
         A     "T_Highpressure_MH02";
         =     "DB123_MH_IO_Signals".MH[2].IN.MH_HP_Circ_MH;
         A     "T_Start_MH02";
         =     "DB123_MH_IO_Signals".MH[2].IN.MH_Start;
         A     "T_Stop_MH02";
         =     "DB123_MH_IO_Signals".MH[2].IN.MH_Stop;
         A     "T_CP_forward_MH02";
         =     "DB123_MH_IO_Signals".MH[2].IN.MH_CP_forward;
         A     "T_CP_back_MH02";
         =     "DB123_MH_IO_Signals".MH[2].IN.MH_CP_backward;
         A     "IPS_MH_MH02";
         =     "DB123_MH_IO_Signals".MH[2].IN.MH_Aps_Mixinghead;

   MHS2: NOP   0;
   //-----------------------------------------------------------------
   // Shot status of MH-02
   //-----------------------------------------------------------------
         L     "PN_Mixinghead".Mixinghead[2].Digital.Address;
         L     0;
         ==D;
         JC    MS02;
         L     "PN_Mixinghead".Mixinghead[2].Digital.Address;
         L     12;
         +D;
         SLD   3;
         LAR1;
         L     PIW [ AR1 , P#0.0 ];
   MS02: T     #TempMHStatus;  // ProCan-MH_Status MH01

         CALL  BLKMOV
         ( SRCBLK  := #TempMHStatus,
           RET_VAL := #TemRetBLKMOV,
           DSTBLK  := "DB123_MH_IO_Signals".MH[2].IN.MH_Status
         );

   //
   //-----------------------------------------------------------------
   // Status of cleaning piston MH-02
   //-----------------------------------------------------------------
         A(;
         L     "PN_Mixinghead".Mixinghead[2].ReinigungskolbenDigital.Address;
         L     0;
         ==D;
         );
         ON    "PN_Mixinghead".Mixinghead[2].ReinigungskolbenDigital.Active;
         JC    CP02;
         L     "PN_Mixinghead".Mixinghead[2].ReinigungskolbenDigital.Address;
         L     8;
         +D;
         SLD   3;
         LAR1;
         L     PIB [ AR1 , P#0.0 ];
   CP02: T     #TempCPStatus;

         CALL  BLKMOV
         ( SRCBLK  := #TempCPStatus,
           RET_VAL := #TemRetBLKMOV,
           DSTBLK  := "DB123_MH_IO_Signals".MH[2].IN.CleaningPistonState
         );

   //-----------------------------------------------------------------
   // Actual shot time of MH-02
   //-----------------------------------------------------------------
         L     "PN_Mixinghead".Mixinghead[2].Digital.Address;
         L     0;
         ==D;
         JC    ST02;

         L     "PN_Mixinghead".Mixinghead[2].Digital.Address;
         SLD   3;
         LAR1;
         L     PID[AR1, P#0.0];
   ST02: T     "DB123_MH_IO_Signals".MH[2].IN.Shottime;

         AN    "DB123_MH_IO_Signals".MH[2].IN.MH_Status.shotdone_MH;
         JC    ShD2;

         L     "PN_Mixinghead".Mixinghead[2].Digital.Address;
         L     4;
         +D;
         SLD   3;
         LAR1;
         L     PID[ AR1 , P#0.0 ];
         T     "DB123_MH_IO_Signals".MH[2].IN.MH_Opentime;

         L     "PN_Mixinghead".Mixinghead[2].Digital.Address;
         L     8;
         +D;
         SLD   3;
         LAR1;
         L     PID [ AR1 , P#0.0 ];
         T     "DB123_MH_IO_Signals".MH[2].IN.MH_Closingtime;
   ShD2: NOP   0;
   emk2: NOP   0;
END_REGION

REGION Network 7: Read ProCan Data of MH-03
   //----------------------------------------------------------------
   // Check if ProfiBus member is accessible and without fault
   // otherwise no communication is possible
   //----------------------------------------------------------------
         A     "PN_Mixinghead".Mixinghead[3].Digital.Active;
         JC    mk3;
         L     0;
         T     #Nullmerker;
         CALL  FILL
         ( BVAL    := #Nullmerker,
           RET_VAL := #ERROR_CODE,
           BLK     := "DB123_MH_IO_Signals".MH[3]
         );
         JU    emk3;
   //_________________________________________________________________
   //
   mk3:  NOP   0;

   //-----------------------------------------------------------------
   // Digital Input -> Ini Signals mixinghead, cleaningpiston
   //-----------------------------------------------------------------
         A     "ES_OP_Panel_MH03";
         =     "DB123_MH_IO_Signals".MH[3].IN.MH_EmergencyStop;
         A     "IPS_CP_MH03";
         =     "DB123_MH_IO_Signals".MH[3].IN.MH_APS_CleaningPiston;
         SET;
         =     "DB123_MH_IO_Signals".MH[3].IN.MH_With_CleaningPiston;
         A     "S_Rel_SWU_MH03";
         =     "DB123_MH_IO_Signals".MH[3].IN.MH_Release_SWU;
         A     "S_Manuel_MH03";
         =     "DB123_MH_IO_Signals".MH[3].IN.MH_Manual_Mode;
         A     "S_Automatic_MH03";
         =     "DB123_MH_IO_Signals".MH[3].IN.MH_Auto_Mode;
         A     "K_PreparationFoamingMC03";
         =     "DB123_MH_IO_Signals".MH[3].IN.MH_Prep_Foaming_MC;
         A     "K_FoamingReleaseMC03";
         =     "DB123_MH_IO_Signals".MH[3].IN.MH_Releas_Foaming_MC;
   //
         L     "S_ProgNoSelectMH03";
         AW    W#16#F;
         T     "DB123_MH_IO_Signals".MH[3].IN.MH_Prog_No_MH;

         A     "T_Highpressure_MH03";
         =     "DB123_MH_IO_Signals".MH[3].IN.MH_HP_Circ_MH;
         A     "T_Start_MH03";
         =     "DB123_MH_IO_Signals".MH[3].IN.MH_Start;
         A     "T_Stop_MH03";
         =     "DB123_MH_IO_Signals".MH[3].IN.MH_Stop;
         A     "T_CP_forward_MH03";
         =     "DB123_MH_IO_Signals".MH[3].IN.MH_CP_forward;
         A     "T_CP_back_MH03";
         =     "DB123_MH_IO_Signals".MH[3].IN.MH_CP_backward;
         A     "IPS_MH_MH03";
         =     "DB123_MH_IO_Signals".MH[3].IN.MH_Aps_Mixinghead;

         NOP   0;
   //-----------------------------------------------------------------
   // Shot status of MH 3
   //-----------------------------------------------------------------
         L     "PN_Mixinghead".Mixinghead[3].Digital.Address;
         L     0;
         ==D;
         JC    MS03;
         L     "PN_Mixinghead".Mixinghead[3].Digital.Address;
         L     12;
         +D;
         SLD   3;
         LAR1;
         L     PIW [ AR1 , P#0.0 ];
   MS03: T     #TempMHStatus;  // ProCan-MH_Status MH03

         CALL  BLKMOV
         ( SRCBLK  := #TempMHStatus,
           RET_VAL := #TemRetBLKMOV,
           DSTBLK  := "DB123_MH_IO_Signals".MH[3].IN.MH_Status
         );
   //
   //-----------------------------------------------------------------
   // Status of cleaning piston MH 3
   //-----------------------------------------------------------------
         A(;
         L     "PN_Mixinghead".Mixinghead[3].ReinigungskolbenDigital.Address;
         L     0;
         ==D;
         );
         ON    "PN_Mixinghead".Mixinghead[3].ReinigungskolbenDigital.Active;
         JC    CP03;
         L     "PN_Mixinghead".Mixinghead[3].ReinigungskolbenDigital.Address;
         L     8;
         +D;
         SLD   3;
         LAR1;
         L     PIB [ AR1 , P#0.0 ];
   CP03: T     #TempCPStatus;

         CALL  BLKMOV
         ( SRCBLK  := #TempCPStatus,
           RET_VAL := #TemRetBLKMOV,
           DSTBLK  := "DB123_MH_IO_Signals".MH[3].IN.CleaningPistonState
         );

   //-----------------------------------------------------------------
   // Actual shot time of mixinghead modul
   //-----------------------------------------------------------------
         L     "PN_Mixinghead".Mixinghead[3].Digital.Address;
         L     0;
         ==D;
         JC    ST03;
   //-
         L     "PN_Mixinghead".Mixinghead[3].Digital.Address;
         SLD   3;
         LAR1;
         L     PID[AR1, P#0.0];
   ST03: T     "DB123_MH_IO_Signals".MH[3].IN.Shottime;
   //-
         AN    "DB123_MH_IO_Signals".MH[3].IN.MH_Status.shotdone_MH;
         JC    ShD3;
   //-
         L     "PN_Mixinghead".Mixinghead[3].Digital.Address;
         L     4;
         +D;
         SLD   3;
         LAR1;
         L     PID[ AR1 , P#0.0 ];
         T     "DB123_MH_IO_Signals".MH[3].IN.MH_Opentime;
   //-
         L     "PN_Mixinghead".Mixinghead[3].Digital.Address;
         L     8;
         +D;
         SLD   3;
         LAR1;
         L     PID [ AR1 , P#0.0 ];
         T     "DB123_MH_IO_Signals".MH[3].IN.MH_Closingtime;
   //-
   ShD3: NOP   0;
   emk3: NOP   0;
END_REGION

REGION Network 8: Read ProCan Data of MH-04
   //----------------------------------------------------------------
   // Check if ProfiBus member is accessible and without fault
   // otherwise no communication is possible
   //----------------------------------------------------------------
         A     "PN_Mixinghead".Mixinghead[4].Digital.Active;
         JC    mk4;
         L     0;
         T     #Nullmerker;
         CALL  FILL
         ( BVAL    := #Nullmerker,
           RET_VAL := #ERROR_CODE,
           BLK     := "DB123_MH_IO_Signals".MH[4]
         );
         JU    emk4;
   //_________________________________________________________________
   //
   mk4:  NOP   0;

   //-----------------------------------------------------------------
   // Digital Input -> Ini Signals mixinghead, cleaningpiston
   //-----------------------------------------------------------------
         A     "ES_OP_Panel_MH04";
         =     "DB123_MH_IO_Signals".MH[4].IN.MH_EmergencyStop;
         A     "IPS_CP_MH04";
         =     "DB123_MH_IO_Signals".MH[4].IN.MH_APS_CleaningPiston;
   //     SET
   //      =     "DB123_MH_IO_Signals".MH[4].IN.MH_With_CleaningPiston
         A     "S_Rel_SWU_MH04";
         =     "DB123_MH_IO_Signals".MH[4].IN.MH_Release_SWU;
         A     "S_Manuel_MH04";
         =     "DB123_MH_IO_Signals".MH[4].IN.MH_Manual_Mode;
         A     "S_Automatic_MH04";
         =     "DB123_MH_IO_Signals".MH[4].IN.MH_Auto_Mode;
         A     "K_PreparationFoamingMC04";
         =     "DB123_MH_IO_Signals".MH[4].IN.MH_Prep_Foaming_MC;
         A     "K_FoamingReleaseMC04";
         =     "DB123_MH_IO_Signals".MH[4].IN.MH_Releas_Foaming_MC;
   ///
         L     "S_ProgNoSelectMH04";
         AW    W#16#F;
         T     "DB123_MH_IO_Signals".MH[4].IN.MH_Prog_No_MH;

         A     "T_Highpressure_MH04";
         =     "DB123_MH_IO_Signals".MH[4].IN.MH_HP_Circ_MH;
         A     "T_Start_MH04";
         =     "DB123_MH_IO_Signals".MH[4].IN.MH_Start;
         A     "T_Stop_MH04";
         =     "DB123_MH_IO_Signals".MH[4].IN.MH_Stop;
         A     "T_CP_forward_MH04";
         =     "DB123_MH_IO_Signals".MH[4].IN.MH_CP_forward;
         A     "T_CP_back_MH04";
         =     "DB123_MH_IO_Signals".MH[4].IN.MH_CP_backward;
         A     "IPS_MH_MH04";
         =     "DB123_MH_IO_Signals".MH[4].IN.MH_Aps_Mixinghead;

         NOP   0;
   //-----------------------------------------------------------------
   // Shot status of MH 4
   //-----------------------------------------------------------------
         L     "PN_Mixinghead".Mixinghead[4].Digital.Address;
         L     0;
         ==D;
         JC    MS04;
         L     "PN_Mixinghead".Mixinghead[4].Digital.Address;
         L     12;
         +D;
         SLD   3;
         LAR1;
         L     PIW [ AR1 , P#0.0 ];
   MS04: T     #TempMHStatus;  // ProCan-MH_Status MH04

         CALL  BLKMOV
         ( SRCBLK  := #TempMHStatus,
           RET_VAL := #TemRetBLKMOV,
           DSTBLK  := "DB123_MH_IO_Signals".MH[4].IN.MH_Status
         );
   //
   //-----------------------------------------------------------------
   // Status of cleaning piston MH 4
   //-----------------------------------------------------------------
         A(;
         L     "PN_Mixinghead".Mixinghead[4].ReinigungskolbenDigital.Address;
         L     0;
         ==D;
         );
         ON    "PN_Mixinghead".Mixinghead[4].ReinigungskolbenDigital.Active;
         JC    CP04;
         L     "PN_Mixinghead".Mixinghead[4].ReinigungskolbenDigital.Address;
         L     8;
         +D;
         SLD   3;
         LAR1;
         L     PIB [ AR1 , P#0.0 ];
   CP04: T     #TempCPStatus;

         CALL  BLKMOV
         ( SRCBLK  := #TempCPStatus,
           RET_VAL := #TemRetBLKMOV,
           DSTBLK  := "DB123_MH_IO_Signals".MH[4].IN.CleaningPistonState
         );

   //-----------------------------------------------------------------
   // Actual shot time of mixinghead modul
   //-----------------------------------------------------------------
         L     "PN_Mixinghead".Mixinghead[4].Digital.Address;
         L     0;
         ==D;
         JC    ST04;
   //-
         L     "PN_Mixinghead".Mixinghead[4].Digital.Address;
         SLD   3;
         LAR1;
         L     PID[AR1, P#0.0];
   ST04: T     "DB123_MH_IO_Signals".MH[4].IN.Shottime;
   //-
         AN    "DB123_MH_IO_Signals".MH[4].IN.MH_Status.shotdone_MH;
         JC    ShD4;
   //-
         L     "PN_Mixinghead".Mixinghead[4].Digital.Address;
         L     4;
         +D;
         SLD   3;
         LAR1;
         L     PID[ AR1 , P#0.0 ];
         T     "DB123_MH_IO_Signals".MH[4].IN.MH_Opentime;
   //-
         L     "PN_Mixinghead".Mixinghead[4].Digital.Address;
         L     8;
         +D;
         SLD   3;
         LAR1;
         L     PID [ AR1 , P#0.0 ];
         T     "DB123_MH_IO_Signals".MH[4].IN.MH_Closingtime;
   //-
   ShD4: NOP   0;
   emk4: NOP   0;
END_REGION

REGION Network 9: Read ProCan Data of MH-05
   //----------------------------------------------------------------
   // Check if ProfiBus member is accessible and without fault
   // otherwise no communication is possible
   //----------------------------------------------------------------
         A     "PN_Mixinghead".Mixinghead[5].Digital.Active;
         JC    mk5;
         L     0;
         T     #Nullmerker;
         CALL  FILL
         ( BVAL    := #Nullmerker,
           RET_VAL := #ERROR_CODE,
           BLK     := "DB123_MH_IO_Signals".MH[5]
         );
         JU    emk5;
   //_________________________________________________________________
   //
   mk5:  NOP   0;
   //-----------------------------------------------------------------
   // Digital Input -> Ini Signals mixinghead, cleaningpiston
   //-----------------------------------------------------------------
         A     "ES_OP_Panel_MH05";
         =     "DB123_MH_IO_Signals".MH[5].IN.MH_EmergencyStop;
         A     "IPS_CP_MH05";
         =     "DB123_MH_IO_Signals".MH[5].IN.MH_APS_CleaningPiston;
   //      SET
   // =     "DB123_MH_IO_Signals".MH[5].IN.MH_With_CleaningPiston
         A     "S_Rel_SWU_MH05";
         =     "DB123_MH_IO_Signals".MH[5].IN.MH_Release_SWU;
         A     "S_Manuel_MH05";
         =     "DB123_MH_IO_Signals".MH[5].IN.MH_Manual_Mode;
         A     "S_Automatic_MH05";
         =     "DB123_MH_IO_Signals".MH[5].IN.MH_Auto_Mode;
         A     "K_PreparationFoamingMC05";
         =     "DB123_MH_IO_Signals".MH[5].IN.MH_Prep_Foaming_MC;
         A     "K_FoamingReleaseMC05";
         =     "DB123_MH_IO_Signals".MH[5].IN.MH_Releas_Foaming_MC;
   ///
         L     "S_ProgNoSelectMH05";
         AW    W#16#F;
         T     "DB123_MH_IO_Signals".MH[5].IN.MH_Prog_No_MH;

         A     "T_Highpressure_MH05";
         =     "DB123_MH_IO_Signals".MH[5].IN.MH_HP_Circ_MH;
         A     "T_Start_MH05";
         =     "DB123_MH_IO_Signals".MH[5].IN.MH_Start;
         A     "T_Stop_MH05";
         =     "DB123_MH_IO_Signals".MH[5].IN.MH_Stop;
         A     "T_CP_forward_MH05";
         =     "DB123_MH_IO_Signals".MH[5].IN.MH_CP_forward;
         A     "T_CP_back_MH05";
         =     "DB123_MH_IO_Signals".MH[5].IN.MH_CP_backward;
         A     "IPS_MH_MH05";
         =     "DB123_MH_IO_Signals".MH[5].IN.MH_Aps_Mixinghead;

         NOP   0;
   //-----------------------------------------------------------------
   // Shot status of MH 5
   //-----------------------------------------------------------------
         L     "PN_Mixinghead".Mixinghead[5].Digital.Address;
         L     0;
         ==D;
         JC    MS05;
         L     "PN_Mixinghead".Mixinghead[5].Digital.Address;
         L     12;
         +D;
         SLD   3;
         LAR1;
         L     PIW [ AR1 , P#0.0 ];
   MS05: T     #TempMHStatus;  // ProCan-MH_Status MH05

         CALL  BLKMOV
         ( SRCBLK  := #TempMHStatus,
           RET_VAL := #TemRetBLKMOV,
           DSTBLK  := "DB123_MH_IO_Signals".MH[5].IN.MH_Status
         );
   //
   //-----------------------------------------------------------------
   // Status of cleaning piston MH 5
   //-----------------------------------------------------------------
         A(;
         L     "PN_Mixinghead".Mixinghead[5].ReinigungskolbenDigital.Address;
         L     0;
         ==D;
         );
         ON    "PN_Mixinghead".Mixinghead[5].ReinigungskolbenDigital.Active;
         JC    CP05;
         L     "PN_Mixinghead".Mixinghead[5].ReinigungskolbenDigital.Address;
         L     8;
         +D;
         SLD   3;
         LAR1;
         L     PIB [ AR1 , P#0.0 ];
   CP05: T     #TempCPStatus;

         CALL  BLKMOV
         ( SRCBLK  := #TempCPStatus,
           RET_VAL := #TemRetBLKMOV,
           DSTBLK  := "DB123_MH_IO_Signals".MH[5].IN.CleaningPistonState
         );

   //-----------------------------------------------------------------
   // Actual shot time of mixinghead modul
   //-----------------------------------------------------------------
         L     "PN_Mixinghead".Mixinghead[5].Digital.Address;
         L     0;
         ==D;
         JC    ST05;
   //-
         L     "PN_Mixinghead".Mixinghead[5].Digital.Address;
         SLD   3;
         LAR1;
         L     PID[AR1, P#0.0];
   ST05: T     "DB123_MH_IO_Signals".MH[5].IN.Shottime;
   //-
         AN    "DB123_MH_IO_Signals".MH[5].IN.MH_Status.shotdone_MH;
         JC    ShD5;
   //-
         L     "PN_Mixinghead".Mixinghead[5].Digital.Address;
         L     4;
         +D;
         SLD   3;
         LAR1;
         L     PID[ AR1 , P#0.0 ];
         T     "DB123_MH_IO_Signals".MH[5].IN.MH_Opentime;
   //-
         L     "PN_Mixinghead".Mixinghead[5].Digital.Address;
         L     8;
         +D;
         SLD   3;
         LAR1;
         L     PID [ AR1 , P#0.0 ];
         T     "DB123_MH_IO_Signals".MH[5].IN.MH_Closingtime;
   //-
   ShD5: NOP   0;
   emk5: NOP   0;
END_REGION

REGION Network 10: Read ProCan Data of MH-06
   //----------------------------------------------------------------
   // Check if ProfiBus member is accessible and without fault
   // otherwise no communication is possible
   //----------------------------------------------------------------
         A     "PN_Mixinghead".Mixinghead[6].Digital.Active;
         JC    mk6;
         L     0;
         T     #Nullmerker;
         CALL  FILL
         ( BVAL    := #Nullmerker,
           RET_VAL := #ERROR_CODE,
           BLK     := "DB123_MH_IO_Signals".MH[6]
         );
         JU    emk6;
   //_________________________________________________________________
   //
   mk6:  NOP   0;

   //-----------------------------------------------------------------
   // Digital Input -> Ini Signals mixinghead, cleaningpiston
   //-----------------------------------------------------------------
         A     "ES_OP_Panel_MH06";
         =     "DB123_MH_IO_Signals".MH[6].IN.MH_EmergencyStop;
         A     "IPS_CP_MH06";
         =     "DB123_MH_IO_Signals".MH[6].IN.MH_APS_CleaningPiston;
   //      SET
   //      =     "DB123_MH_IO_Signals".MH[6].IN.MH_With_CleaningPiston
         A     "S_Rel_SWU_MH06";
         =     "DB123_MH_IO_Signals".MH[6].IN.MH_Release_SWU;
         A     "S_Manuel_MH06";
         =     "DB123_MH_IO_Signals".MH[6].IN.MH_Manual_Mode;
         A     "S_Automatic_MH06";
         =     "DB123_MH_IO_Signals".MH[6].IN.MH_Auto_Mode;
         A     "K_PreparationFoamingMC06";
         =     "DB123_MH_IO_Signals".MH[6].IN.MH_Prep_Foaming_MC;
         A     "K_FoamingReleaseMC06";
         =     "DB123_MH_IO_Signals".MH[6].IN.MH_Releas_Foaming_MC;
   ///
         L     "S_ProgNoSelectMH06";
         AW    W#16#F;
         T     "DB123_MH_IO_Signals".MH[6].IN.MH_Prog_No_MH;

         A     "T_Highpressure_MH06";
         =     "DB123_MH_IO_Signals".MH[6].IN.MH_HP_Circ_MH;
         A     "T_Start_MH06";
         =     "DB123_MH_IO_Signals".MH[6].IN.MH_Start;
         A     "T_Stop_MH06";
         =     "DB123_MH_IO_Signals".MH[6].IN.MH_Stop;
         A     "T_CP_forward_MH06";
         =     "DB123_MH_IO_Signals".MH[6].IN.MH_CP_forward;
         A     "T_CP_back_MH06";
         =     "DB123_MH_IO_Signals".MH[6].IN.MH_CP_backward;
         A     "IPS_MH_MH06";
         =     "DB123_MH_IO_Signals".MH[6].IN.MH_Aps_Mixinghead;

         NOP   0;
   //-----------------------------------------------------------------
   // Shot status of MH 6
   //-----------------------------------------------------------------
         L     "PN_Mixinghead".Mixinghead[6].Digital.Address;
         L     0;
         ==D;
         JC    MS06;
         L     "PN_Mixinghead".Mixinghead[6].Digital.Address;
         L     12;
         +D;
         SLD   3;
         LAR1;
         L     PIW [ AR1 , P#0.0 ];
   MS06: T     #TempMHStatus;  // ProCan-MH_Status MH06

         CALL  BLKMOV
         ( SRCBLK  := #TempMHStatus,
           RET_VAL := #TemRetBLKMOV,
           DSTBLK  := "DB123_MH_IO_Signals".MH[6].IN.MH_Status
         );
   //
   //-----------------------------------------------------------------
   // Status of cleaning piston MH 6
   //-----------------------------------------------------------------
         A(;
         L     "PN_Mixinghead".Mixinghead[6].ReinigungskolbenDigital.Address;
         L     0;
         ==D;
         );
         ON    "PN_Mixinghead".Mixinghead[6].ReinigungskolbenDigital.Active;
         JC    CP06;
         L     "PN_Mixinghead".Mixinghead[6].ReinigungskolbenDigital.Address;
         L     8;
         +D;
         SLD   3;
         LAR1;
         L     PIB [ AR1 , P#0.0 ];
   CP06: T     #TempCPStatus;

         CALL  BLKMOV
         ( SRCBLK  := #TempCPStatus,
           RET_VAL := #TemRetBLKMOV,
           DSTBLK  := "DB123_MH_IO_Signals".MH[6].IN.CleaningPistonState
         );

   //-----------------------------------------------------------------
   // Actual shot time of mixinghead modul
   //-----------------------------------------------------------------
         L     "PN_Mixinghead".Mixinghead[6].Digital.Address;
         L     0;
         ==D;
         JC    ST06;
   //-
         L     "PN_Mixinghead".Mixinghead[6].Digital.Address;
         SLD   3;
         LAR1;
         L     PID[AR1, P#0.0];
   ST06: T     "DB123_MH_IO_Signals".MH[6].IN.Shottime;
   //-
         AN    "DB123_MH_IO_Signals".MH[6].IN.MH_Status.shotdone_MH;
         JC    ShD6;
   //-
         L     "PN_Mixinghead".Mixinghead[6].Digital.Address;
         L     4;
         +D;
         SLD   3;
         LAR1;
         L     PID[ AR1 , P#0.0 ];
         T     "DB123_MH_IO_Signals".MH[6].IN.MH_Opentime;
   //-
         L     "PN_Mixinghead".Mixinghead[6].Digital.Address;
         L     8;
         +D;
         SLD   3;
         LAR1;
         L     PID [ AR1 , P#0.0 ];
         T     "DB123_MH_IO_Signals".MH[6].IN.MH_Closingtime;
   //-
   ShD6: NOP   0;
   emk6: NOP   0;
END_REGION

REGION Network 11: Read ProCan Data of MH-07
   //----------------------------------------------------------------
   // Check if ProfiBus member is accessible and without fault
   // otherwise no communication is possible
   //----------------------------------------------------------------
         A     "PN_Mixinghead".Mixinghead[7].Digital.Active;
         JC    mk7;
         L     0;
         T     #Nullmerker;
         CALL  FILL
         ( BVAL    := #Nullmerker,
           RET_VAL := #ERROR_CODE,
           BLK     := "DB123_MH_IO_Signals".MH[7]
         );
         JU    emk7;
   //_________________________________________________________________
   //
   mk7:  NOP   0;

   //-----------------------------------------------------------------
   // Digital Input -> Ini Signals mixinghead, cleaningpiston
   //-----------------------------------------------------------------
         A     "ES_OP_Panel_MH07";
         =     "DB123_MH_IO_Signals".MH[7].IN.MH_EmergencyStop;
         A     "IPS_CP_MH07";
         =     "DB123_MH_IO_Signals".MH[7].IN.MH_APS_CleaningPiston;
   //      SET
   //      =     "DB123_MH_IO_Signals".MH[7].IN.MH_With_CleaningPiston
         A     "S_Rel_SWU_MH07";
         =     "DB123_MH_IO_Signals".MH[7].IN.MH_Release_SWU;
         A     "S_Manuel_MH07";
         =     "DB123_MH_IO_Signals".MH[7].IN.MH_Manual_Mode;
         A     "S_Automatic_MH07";
         =     "DB123_MH_IO_Signals".MH[7].IN.MH_Auto_Mode;
         A     "K_PreparationFoamingMC07";
         =     "DB123_MH_IO_Signals".MH[7].IN.MH_Prep_Foaming_MC;
         A     "K_FoamingReleaseMC07";
         =     "DB123_MH_IO_Signals".MH[7].IN.MH_Releas_Foaming_MC;
   ///
         L     "S_ProgNoSelectMH07";
         AW    W#16#F;
         T     "DB123_MH_IO_Signals".MH[7].IN.MH_Prog_No_MH;

         A     "T_Highpressure_MH07";
         =     "DB123_MH_IO_Signals".MH[7].IN.MH_HP_Circ_MH;
         A     "T_Start_MH07";
         =     "DB123_MH_IO_Signals".MH[7].IN.MH_Start;
         A     "T_Stop_MH07";
         =     "DB123_MH_IO_Signals".MH[7].IN.MH_Stop;
         A     "T_CP_forward_MH07";
         =     "DB123_MH_IO_Signals".MH[7].IN.MH_CP_forward;
         A     "T_CP_back_MH07";
         =     "DB123_MH_IO_Signals".MH[7].IN.MH_CP_backward;
         A     "IPS_MH_MH07";
         =     "DB123_MH_IO_Signals".MH[7].IN.MH_Aps_Mixinghead;

         NOP   0;
   //-----------------------------------------------------------------
   // Shot status of MH 7
   //-----------------------------------------------------------------
         L     "PN_Mixinghead".Mixinghead[7].Digital.Address;
         L     0;
         ==D;
         JC    MS07;
         L     "PN_Mixinghead".Mixinghead[7].Digital.Address;
         L     12;
         +D;
         SLD   3;
         LAR1;
         L     PIW [ AR1 , P#0.0 ];
   MS07: T     #TempMHStatus;  // ProCan-MH_Status MH06

         CALL  BLKMOV
         ( SRCBLK  := #TempMHStatus,
           RET_VAL := #TemRetBLKMOV,
           DSTBLK  := "DB123_MH_IO_Signals".MH[7].IN.MH_Status
         );
   //
   //-----------------------------------------------------------------
   // Status of cleaning piston MH 7
   //-----------------------------------------------------------------
         A(;
         L     "PN_Mixinghead".Mixinghead[7].ReinigungskolbenDigital.Address;
         L     0;
         ==D;
         );
         ON    "PN_Mixinghead".Mixinghead[7].ReinigungskolbenDigital.Active;
         JC    CP07;
         L     "PN_Mixinghead".Mixinghead[7].ReinigungskolbenDigital.Address;
         L     8;
         +D;
         SLD   3;
         LAR1;
         L     PIB [ AR1 , P#0.0 ];
   CP07: T     #TempCPStatus;

         CALL  BLKMOV
         ( SRCBLK  := #TempCPStatus,
           RET_VAL := #TemRetBLKMOV,
           DSTBLK  := "DB123_MH_IO_Signals".MH[7].IN.CleaningPistonState
         );

   //-----------------------------------------------------------------
   // Actual shot time of mixinghead modul
   //-----------------------------------------------------------------
         L     "PN_Mixinghead".Mixinghead[7].Digital.Address;
         L     0;
         ==D;
         JC    ST07;
   //-
         L     "PN_Mixinghead".Mixinghead[7].Digital.Address;
         SLD   3;
         LAR1;
         L     PID[AR1, P#0.0];
   ST07: T     "DB123_MH_IO_Signals".MH[7].IN.Shottime;
   //-
         AN    "DB123_MH_IO_Signals".MH[7].IN.MH_Status.shotdone_MH;
         JC    ShD7;
   //-
         L     "PN_Mixinghead".Mixinghead[7].Digital.Address;
         L     4;
         +D;
         SLD   3;
         LAR1;
         L     PID[ AR1 , P#0.0 ];
         T     "DB123_MH_IO_Signals".MH[7].IN.MH_Opentime;
   //-
         L     "PN_Mixinghead".Mixinghead[7].Digital.Address;
         L     8;
         +D;
         SLD   3;
         LAR1;
         L     PID [ AR1 , P#0.0 ];
         T     "DB123_MH_IO_Signals".MH[7].IN.MH_Closingtime;
   //-
   ShD7: NOP   0;
   emk7: NOP   0;
END_REGION

REGION Network 12: Read ProCan Data of MH-08
   //----------------------------------------------------------------
   // Check if ProfiBus member is accessible and without fault
   // otherwise no communication is possible
   //----------------------------------------------------------------
         A     "PN_Mixinghead".Mixinghead[8].Digital.Active;
         JC    mk8;
         L     0;
         T     #Nullmerker;
         CALL  FILL
         ( BVAL    := #Nullmerker,
           RET_VAL := #ERROR_CODE,
           BLK     := "DB123_MH_IO_Signals".MH[8]
         );
         JU    emk8;
   //_________________________________________________________________
   //
   mk8:  NOP   0;

   //-----------------------------------------------------------------
   // Digital Input -> Ini Signals mixinghead, cleaningpiston
   //-----------------------------------------------------------------
         A     "ES_OP_Panel_MH08";
         =     "DB123_MH_IO_Signals".MH[8].IN.MH_EmergencyStop;
         A     "IPS_CP_MH08";
         =     "DB123_MH_IO_Signals".MH[8].IN.MH_APS_CleaningPiston;
   //      SET
   //      =     "DB123_MH_IO_Signals".MH[8].IN.MH_With_CleaningPiston
         A     "S_Rel_SWU_MH08";
         =     "DB123_MH_IO_Signals".MH[8].IN.MH_Release_SWU;
         A     "S_Manuel_MH08";
         =     "DB123_MH_IO_Signals".MH[8].IN.MH_Manual_Mode;
         A     "S_Automatic_MH08";
         =     "DB123_MH_IO_Signals".MH[8].IN.MH_Auto_Mode;
         A     "K_PreparationFoamingMC08";
         =     "DB123_MH_IO_Signals".MH[8].IN.MH_Prep_Foaming_MC;
         A     "K_FoamingReleaseMC08";
         =     "DB123_MH_IO_Signals".MH[8].IN.MH_Releas_Foaming_MC;
   ///
         L     "S_ProgNoSelectMH08";
         AW    W#16#F;
         T     "DB123_MH_IO_Signals".MH[8].IN.MH_Prog_No_MH;

         A     "T_Highpressure_MH08";
         =     "DB123_MH_IO_Signals".MH[8].IN.MH_HP_Circ_MH;
         A     "T_Start_MH08";
         =     "DB123_MH_IO_Signals".MH[8].IN.MH_Start;
         A     "T_Stop_MH08";
         =     "DB123_MH_IO_Signals".MH[8].IN.MH_Stop;
         A     "T_CP_forward_MH08";
         =     "DB123_MH_IO_Signals".MH[8].IN.MH_CP_forward;
         A     "T_CP_back_MH08";
         =     "DB123_MH_IO_Signals".MH[8].IN.MH_CP_backward;
         A     "IPS_MH_MH08";
         =     "DB123_MH_IO_Signals".MH[8].IN.MH_Aps_Mixinghead;

         NOP   0;
   //-----------------------------------------------------------------
   // Shot status of MH 8
   //-----------------------------------------------------------------
         L     "PN_Mixinghead".Mixinghead[8].Digital.Address;
         L     0;
         ==D;
         JC    MS08;
         L     "PN_Mixinghead".Mixinghead[8].Digital.Address;
         L     12;
         +D;
         SLD   3;
         LAR1;
         L     PIW [ AR1 , P#0.0 ];
   MS08: T     #TempMHStatus;  // ProCan-MH_Status MH06

         CALL  BLKMOV
         ( SRCBLK  := #TempMHStatus,
           RET_VAL := #TemRetBLKMOV,
           DSTBLK  := "DB123_MH_IO_Signals".MH[8].IN.MH_Status
         );
   //
   //-----------------------------------------------------------------
   // Status of cleaning piston MH 8
   //-----------------------------------------------------------------
         A(;
         L     "PN_Mixinghead".Mixinghead[8].ReinigungskolbenDigital.Address;
         L     0;
         ==D;
         );
         ON    "PN_Mixinghead".Mixinghead[8].ReinigungskolbenDigital.Active;
         JC    CP08;
         L     "PN_Mixinghead".Mixinghead[8].ReinigungskolbenDigital.Address;
         L     8;
         +D;
         SLD   3;
         LAR1;
         L     PIB [ AR1 , P#0.0 ];
   CP08: T     #TempCPStatus;

         CALL  BLKMOV
         ( SRCBLK  := #TempCPStatus,
           RET_VAL := #TemRetBLKMOV,
           DSTBLK  := "DB123_MH_IO_Signals".MH[8].IN.CleaningPistonState
         );

   //-----------------------------------------------------------------
   // Actual shot time of mixinghead modul
   //-----------------------------------------------------------------
         L     "PN_Mixinghead".Mixinghead[8].Digital.Address;
         L     0;
         ==D;
         JC    ST08;
   //-
         L     "PN_Mixinghead".Mixinghead[8].Digital.Address;
         SLD   3;
         LAR1;
         L     PID[AR1, P#0.0];
   ST08: T     "DB123_MH_IO_Signals".MH[8].IN.Shottime;
   //-
         AN    "DB123_MH_IO_Signals".MH[8].IN.MH_Status.shotdone_MH;
         JC    ShD8;
   //-
         L     "PN_Mixinghead".Mixinghead[8].Digital.Address;
         L     4;
         +D;
         SLD   3;
         LAR1;
         L     PID[ AR1 , P#0.0 ];
         T     "DB123_MH_IO_Signals".MH[8].IN.MH_Opentime;
   //-
         L     "PN_Mixinghead".Mixinghead[8].Digital.Address;
         L     8;
         +D;
         SLD   3;
         LAR1;
         L     PID [ AR1 , P#0.0 ];
         T     "DB123_MH_IO_Signals".MH[8].IN.MH_Closingtime;
   //-
   ShD8: NOP   0;
   emk8: NOP   0;
END_REGION

REGION Network 13: Read ProCan Data of MH-09
   //----------------------------------------------------------------
   // Check if ProfiBus member is accessible and without fault
   // otherwise no communication is possible
   //----------------------------------------------------------------
         A     "PN_Mixinghead".Mixinghead[9].Digital.Active;
         JC    mk09;
         L     0;
         T     #Nullmerker;
         CALL  FILL
         ( BVAL    := #Nullmerker,
           RET_VAL := #ERROR_CODE,
           BLK     := "DB123_MH_IO_Signals".MH[09]
         );
         JU    emk09;
   //_________________________________________________________________
   //
   mk09: NOP   0;

   //-----------------------------------------------------------------
   // Digital Input -> Ini Signals mixinghead, cleaningpiston
   //-----------------------------------------------------------------
         A     "ES_OP_Panel_MH09";
         =     "DB123_MH_IO_Signals".MH[09].IN.MH_EmergencyStop;
         A     "IPS_CP_MH09";
         =     "DB123_MH_IO_Signals".MH[09].IN.MH_APS_CleaningPiston;
   //      SET
   //      =     "DB123_MH_IO_Signals".MH[09].IN.MH_With_CleaningPiston
         A     "S_Rel_SWU_MH09";
         =     "DB123_MH_IO_Signals".MH[09].IN.MH_Release_SWU;
         A     "S_Manuel_MH09";
         =     "DB123_MH_IO_Signals".MH[09].IN.MH_Manual_Mode;
         A     "S_Automatic_MH09";
         =     "DB123_MH_IO_Signals".MH[09].IN.MH_Auto_Mode;
         A     "K_PreparationFoamingMC09";
         =     "DB123_MH_IO_Signals".MH[09].IN.MH_Prep_Foaming_MC;
         A     "K_FoamingReleaseMC09";
         =     "DB123_MH_IO_Signals".MH[09].IN.MH_Releas_Foaming_MC;
   ///
         L     "S_ProgNoSelectMH09";
         AW    W#16#F;
         T     "DB123_MH_IO_Signals".MH[09].IN.MH_Prog_No_MH;

         A     "T_Highpressure_MH09";
         =     "DB123_MH_IO_Signals".MH[09].IN.MH_HP_Circ_MH;
         A     "T_Start_MH09";
         =     "DB123_MH_IO_Signals".MH[09].IN.MH_Start;
         A     "T_Stop_MH09";
         =     "DB123_MH_IO_Signals".MH[09].IN.MH_Stop;
         A     "T_CP_forward_MH09";
         =     "DB123_MH_IO_Signals".MH[09].IN.MH_CP_forward;
         A     "T_CP_back_MH09";
         =     "DB123_MH_IO_Signals".MH[09].IN.MH_CP_backward;
         A     "IPS_MH_MH09";
         =     "DB123_MH_IO_Signals".MH[09].IN.MH_Aps_Mixinghead;

         NOP   0;
   //-----------------------------------------------------------------
   // Shot status of MH 09
   //-----------------------------------------------------------------
         L     "PN_Mixinghead".Mixinghead[9].Digital.Address;
         L     0;
         ==D;
         JC    MS09;
         L     "PN_Mixinghead".Mixinghead[9].Digital.Address;
         L     12;
         +D;
         SLD   3;
         LAR1;
         L     PIW [ AR1 , P#0.0 ];
   MS09: T     #TempMHStatus;  // ProCan-MH_Status MH09

         CALL  BLKMOV
         ( SRCBLK  := #TempMHStatus,
           RET_VAL := #TemRetBLKMOV,
           DSTBLK  := "DB123_MH_IO_Signals".MH[09].IN.MH_Status
         );
   //
   //-----------------------------------------------------------------
   // Status of cleaning piston MH 09
   //-----------------------------------------------------------------
         A(;
         L     "PN_Mixinghead".Mixinghead[9].ReinigungskolbenDigital.Address;
         L     0;
         ==D;
         );
         ON    "PN_Mixinghead".Mixinghead[9].ReinigungskolbenDigital.Active;
         JC    CP09;
         L     "PN_Mixinghead".Mixinghead[9].ReinigungskolbenDigital.Address;
         L     8;
         +D;
         SLD   3;
         LAR1;
         L     PIB [ AR1 , P#0.0 ];
   CP09: T     #TempCPStatus;

         CALL  BLKMOV
         ( SRCBLK  := #TempCPStatus,
           RET_VAL := #TemRetBLKMOV,
           DSTBLK  := "DB123_MH_IO_Signals".MH[09].IN.CleaningPistonState
         );

   //-----------------------------------------------------------------
   // Actual shot time of mixinghead modul
   //-----------------------------------------------------------------
         L     "PN_Mixinghead".Mixinghead[9].Digital.Address;
         L     0;
         ==D;
         JC    ST09;
   //-
         L     "PN_Mixinghead".Mixinghead[9].Digital.Address;
         SLD   3;
         LAR1;
         L     PID[AR1, P#0.0];
   ST09: T     "DB123_MH_IO_Signals".MH[9].IN.Shottime;
   //-
         AN    "DB123_MH_IO_Signals".MH[9].IN.MH_Status.shotdone_MH;
         JC    ShD9;
   //-
         L     "PN_Mixinghead".Mixinghead[9].Digital.Address;
         L     4;
         +D;
         SLD   3;
         LAR1;
         L     PID[ AR1 , P#0.0 ];
         T     "DB123_MH_IO_Signals".MH[9].IN.MH_Opentime;
   //-
         L     "PN_Mixinghead".Mixinghead[9].Digital.Address;
         L     8;
         +D;
         SLD   3;
         LAR1;
         L     PID [ AR1 , P#0.0 ];
         T     "DB123_MH_IO_Signals".MH[9].IN.MH_Closingtime;
   //-
   ShD9: NOP   0;
   emk09:NOP   0;
END_REGION

REGION Network 14: Read ProCan Data of MH-10
   //----------------------------------------------------------------
   // Check if ProfiBus member is accessible and without fault
   // otherwise no communication is possible
   //----------------------------------------------------------------
         A     "PN_Mixinghead".Mixinghead[10].Digital.Active;
         JC    mk10;
         L     0;
         T     #Nullmerker;
         CALL  FILL
         ( BVAL    := #Nullmerker,
           RET_VAL := #ERROR_CODE,
           BLK     := "DB123_MH_IO_Signals".MH[10]
         );
         JU    emk10;
   //_________________________________________________________________
   //
   mk10: NOP   0;

   //-----------------------------------------------------------------
   // Digital Input -> Ini Signals mixinghead, cleaningpiston
   //-----------------------------------------------------------------
         A     "ES_OP_Panel_MH10";
         =     "DB123_MH_IO_Signals".MH[10].IN.MH_EmergencyStop;
         A     "IPS_CP_MH10";
         =     "DB123_MH_IO_Signals".MH[10].IN.MH_APS_CleaningPiston;
   //      SET
   //      =     "DB123_MH_IO_Signals".MH[10].IN.MH_With_CleaningPiston
         A     "S_Rel_SWU_MH10";
         =     "DB123_MH_IO_Signals".MH[10].IN.MH_Release_SWU;
         A     "S_Manuel_MH10";
         =     "DB123_MH_IO_Signals".MH[10].IN.MH_Manual_Mode;
         A     "S_Automatic_MH10";
         =     "DB123_MH_IO_Signals".MH[10].IN.MH_Auto_Mode;
         A     "K_PreparationFoamingMC10";
         =     "DB123_MH_IO_Signals".MH[10].IN.MH_Prep_Foaming_MC;
         A     "K_FoamingReleaseMC10";
         =     "DB123_MH_IO_Signals".MH[10].IN.MH_Releas_Foaming_MC;
   ///
         L     "S_ProgNoSelectMH10";
         AW    W#16#F;
         T     "DB123_MH_IO_Signals".MH[10].IN.MH_Prog_No_MH;

         A     "T_Highpressure_MH10";
         =     "DB123_MH_IO_Signals".MH[10].IN.MH_HP_Circ_MH;
         A     "T_Start_MH10";
         =     "DB123_MH_IO_Signals".MH[10].IN.MH_Start;
         A     "T_Stop_MH10";
         =     "DB123_MH_IO_Signals".MH[10].IN.MH_Stop;
         A     "T_CP_forward_MH10";
         =     "DB123_MH_IO_Signals".MH[10].IN.MH_CP_forward;
         A     "T_CP_back_MH10";
         =     "DB123_MH_IO_Signals".MH[10].IN.MH_CP_backward;
         A     "IPS_MH_MH10";
         =     "DB123_MH_IO_Signals".MH[10].IN.MH_Aps_Mixinghead;

         NOP   0;
   //-----------------------------------------------------------------
   // Shot status of MH 10
   //-----------------------------------------------------------------
         L     "PN_Mixinghead".Mixinghead[10].Digital.Address;
         L     0;
         ==D;
         JC    MS10;
         L     "PN_Mixinghead".Mixinghead[10].Digital.Address;
         L     12;
         +D;
         SLD   3;
         LAR1;
         L     PIW [ AR1 , P#0.0 ];
   MS10: T     #TempMHStatus;  // ProCan-MH_Status MH10

         CALL  BLKMOV
         ( SRCBLK  := #TempMHStatus,
           RET_VAL := #TemRetBLKMOV,
           DSTBLK  := "DB123_MH_IO_Signals".MH[10].IN.MH_Status
         );
   //
   //-----------------------------------------------------------------
   // Status of cleaning piston MH 10
   //-----------------------------------------------------------------
         A(;
         L     "PN_Mixinghead".Mixinghead[10].ReinigungskolbenDigital.Address;
         L     0;
         ==D;
         );
         ON    "PN_Mixinghead".Mixinghead[10].ReinigungskolbenDigital.Active;
         JC    CP10;
         L     "PN_Mixinghead".Mixinghead[10].ReinigungskolbenDigital.Address;
         L     8;
         +D;
         SLD   3;
         LAR1;
         L     PIB [ AR1 , P#0.0 ];
   CP10: T     #TempCPStatus;

         CALL  BLKMOV
         ( SRCBLK  := #TempCPStatus,
           RET_VAL := #TemRetBLKMOV,
           DSTBLK  := "DB123_MH_IO_Signals".MH[10].IN.CleaningPistonState
         );

   //-----------------------------------------------------------------
   // Actual shot time of mixinghead modul
   //-----------------------------------------------------------------
         L     "PN_Mixinghead".Mixinghead[10].Digital.Address;
         L     0;
         ==D;
         JC    ST10;
   //-
         L     "PN_Mixinghead".Mixinghead[10].Digital.Address;
         SLD   3;
         LAR1;
         L     PID[AR1, P#0.0];
   ST10: T     "DB123_MH_IO_Signals".MH[10].IN.Shottime;
   //-
         AN    "DB123_MH_IO_Signals".MH[10].IN.MH_Status.shotdone_MH;
         JC    ShD10;  //-
         L     "PN_Mixinghead".Mixinghead[10].Digital.Address;
         L     4;
         +D;
         SLD   3;
         LAR1;
         L     PID[ AR1 , P#0.0 ];
         T     "DB123_MH_IO_Signals".MH[10].IN.MH_Opentime;
   //-
         L     "PN_Mixinghead".Mixinghead[10].Digital.Address;
         L     8;
         +D;
         SLD   3;
         LAR1;
         L     PID [ AR1 , P#0.0 ];
         T     "DB123_MH_IO_Signals".MH[10].IN.MH_Closingtime;
   //-
   ShD10:NOP   0;
   emk10:NOP   0;
END_REGION
END_FUNCTION

FUNCTION "FC121_Aggitator" : Void   // FC121, STL
TITLE = Control of several auxiliary drives of a pouring machine
{ S7_Optimized_Access := 'FALSE' }
AUTHOR : KT242
FAMILY : RS_KK
NAME : Drive
VERSION : 1.5
   VAR_INPUT
      IN_Release : Bool;   // Genarelly release 0f the drive (Operation mode)
      IN_ControlVoltage : Bool;   // Signal delay activation frequency converter (protection after emergency-stop)
      IN_Reset_fault : Bool;   // Signal to quit fault within function block
      IN_Request_Filling : Bool;   // Request switch on drive for filling
      IN_Request_Feed : Bool;   // Request switch on drive if componenten pump start up
      IN_Request_Cooling : Bool;   // Request switch on drive for cooling
      IN_Request_Heating : Bool;   // Request switch on drive for heating
      IN_Fault_Motorprotection : Bool;   // Input fault motorprotection of drive
      IN_FaultFreqConverter : Bool;   // Input fault frequency converter of drive
      IN_MaxLevelTray : Bool;   // Input fault max. filling level tray
      IN_EnableLevel : Bool;   // Input Level for enable agitator
      IN_TimerDrive : Timer;   // Timer of general timing of the drive
      IN_TimerStartUpFConv : Timer;   // Timer of delay start up frequency converter
      IN_Values : "UDT710_Agitator";   // Values of configuration
   END_VAR
   VAR_OUTPUT
      OUT_MainsContactor : Bool;   // Ouput mainscontactor drive or frequency converter
      OUT_Release_FConverter : Bool;   // Output release of frequncy converter to control rotation speed
   END_VAR
   VAR_IN_OUT
      IO_Status : ANY;   // Stores the state of the drive
      IO_NewFault : Bool;
      IO_FaultLevel_3 : Bool;
      IO_Faults : ANY;
   END_VAR
   VAR_TEMP
      Temp_IO_Status : "UDT100_AggitatorState";
      ERROR_CODE : Int;   // Error state of systemfunction "BLKMOV" Blockmove
      Anyzeiger1 : ANY;   // Pointer to copy thr array "IO_Status" and "Temp_IO_Status"
      Anyzeiger2 : ANY;   // Pointer to copy thr array "IO_Status" and "Temp_IO_Status"
      Temp_IO_Fault : "UDT1801_Agitator";
      Temp_RunTime : S5Time;   // Flag runtime drive
      Temp_PauseTime : S5Time;   // Flag pause time
      Temp_Runtime_ms : Time;   // Flag runtime drive in millisecond
      Temp_Pausetime_ms : Time;   // Flag pause time drive in millisecond
      Temp_ReleaseDrive : Bool;   // Flag release activation drive
      Temp_WrongTimevalue : Bool;
      Temp_Out_MainsContactor : Bool;
      Temp_Release_FConverter : Bool;
   END_VAR
BEGIN

REGION Network 1: Saved data integration
   // Änderungen:
   // -------------------------------------------------------------------------------
   // Bei der Verwendung der Umwälzpumpe als Speisepumpe wurde dieses bei Min. 
   // Füllstand ausgeshaltet, auch wenn dies im Zyklus auftrat. Hierdurch wurden dann 
   // auch die Materialpumpen abgeschaltet.
   // v.d.Geest     25.02.2003
   // -------------------------------------------------------------------------------
   // Bei einer Ansteuerung mit Frequenzumrichter wurde nicht auf die 
   // Störungsauswertung des Umrichters gewartet bevor die Freigabe gegeben wurde. 
   // Hierdurch kam es zu Störungen bei jedem einschalten des Aggregates.
   // A. Jäger      21.11.2003
   //-----
         LAR1;
         L;
         LAR2;
   //-----
         L     W[AR2, P#0.0];  // Bytes
         T     W[AR1, P#0.0];
         L     W[AR2, P#2.0];  // Amount of bytes
         T     W[AR1, P#2.0];
         L     W[AR2, P#4.0];  // Block no,
         T     W[AR1, P#4.0];
         L     D[AR2, P#6.0];  // Startadress of datas
         T     D[AR1, P#6.0];
   //-----
         CALL  BLKMOV
         ( SRCBLK  := #Anyzeiger1,
           RET_VAL := #ERROR_CODE,
           DSTBLK  := #Temp_IO_Status
         );
   //-----
         LAR1;
         L;
         LAR2;
   //-----
         L     W[AR2, P#0.0];  // Bytes
         T     W[AR1, P#0.0];
         L     W[AR2, P#2.0];  // Amount of bytes
         T     W[AR1, P#2.0];
         L     W[AR2, P#4.0];  // Block no,
         T     W[AR1, P#4.0];
         L     D[AR2, P#6.0];  // Startadress of datas
         T     D[AR1, P#6.0];
   //-----
         CALL  BLKMOV
         ( SRCBLK  := #Anyzeiger2,
           RET_VAL := #ERROR_CODE,
           DSTBLK  := #Temp_IO_Fault
         );
   //-----
END_REGION

REGION Network 2: Release drive
   //-----
         O(;
         A     #IN_Request_Filling;
         A     #IN_Values.Config_bit_Filling_ON;
         );
         O(;
         A     #IN_Request_Feed;
         A     #IN_Values.Config_bit_Charging_ON;
         );
         O(;
         A     #IN_Request_Cooling;
         A     #IN_Values.Config_bit_Cooling_ON;
         );
         O(;
         A     #IN_Request_Heating;
         A     #IN_Values.Config_bit_Heating_ON;
         );
         O     #Temp_IO_Status.Switch_Drive_ON_OFF;
         A     #IN_Release;
         =     #Temp_ReleaseDrive;
END_REGION

REGION Network 3: Faults
   //-----
         A     #IN_Reset_fault;
         R     #Temp_IO_Fault.FLT_Motorprotection;
         R     #Temp_IO_Fault.FLT_FrequencyConverter;
         R     #Temp_IO_Fault.FLT_MaxLTripTray;
         R     #Temp_IO_Fault.FLT_wrong_Timevalue;
         R     #Temp_IO_Fault.Mes_Min_Level;
   //-----
         A     #IN_Fault_Motorprotection;
         AN    #Temp_IO_Fault.FLT_Motorprotection;
         S     #Temp_IO_Fault.FLT_Motorprotection;
         S     #IO_NewFault;
   //-----
         A     #IN_ControlVoltage;
         AN    #Temp_IO_Fault.FLT_wrong_Timevalue;
         AN    #Temp_IO_Status.Start_Startupdelay;
         L     S5T#5S;
         SD    #IN_TimerStartUpFConv;
   //-
         A     #IN_TimerStartUpFConv;
         AN    #IN_FaultFreqConverter;
         A     #Temp_ReleaseDrive;
         A     #IN_Values.Config_bit_Converter;
         AN    #Temp_IO_Fault.FLT_FrequencyConverter;
         S     #Temp_IO_Fault.FLT_FrequencyConverter;
         S     #IO_NewFault;
   //-----
         AN    #IN_MaxLevelTray;
         A     #Temp_ReleaseDrive;
         AN    #Temp_IO_Fault.FLT_MaxLTripTray;
         S     #Temp_IO_Fault.FLT_MaxLTripTray;
         S     #IO_NewFault;
   //-----
         AN    #IN_EnableLevel;
         A     #Temp_ReleaseDrive;
         AN    #Temp_IO_Fault.Mes_Min_Level;
         S     #Temp_IO_Fault.Mes_Min_Level;
         S     #IO_NewFault;
   //-----
END_REGION

